// TIA Portal project "XSFW_TIA32701_A8" (V15.1)

(* hardware
DEVICE "S7-1200 station_1"  S7-1200 Station
   slot 0: "Rack_0"  S7-1200 Rack  Rack  V1.0
   slot 1: "PLC_1"  CPU 1212C DC/DC/DC  6ES7 212-1AE40-0XB0  V4.2
   slot 2: "DI 16/DQ 16x24VDC_1"  6ES7 223-1BL32-0XB0  V2.0
DEVICE "HMI_1"  KTP700 Basic PN
   slot 0: "HMI_1"  KTP700 Basic PN  6AV2 123-2GB03-0AX0  15.0.0.0
   slot 1: "HMI_RT_1"  KTP700 Basic PN  6AV2 123-2GB03-0AX0  15.0.0.0
   slot 5: "HMI_1.IE_CP_1"  PROFINET Interface  15.0.0.0
      slot 1: "Interfaz PROFINET_1"  PROFINET Interface
         slot 1: "Port_1"  Port
*)

// ===== PLC "PLC_1"  CPU 1212C DC/DC/DC =====

VAR_GLOBAL   // PLC tag table "Tabla de variables estándar"
   "Tag_2" AT %M101.0 : Bool;
   "Clock_Byte" AT %MB0 : Byte;
   "Clock_10Hz" AT %M0.0 : Bool;
   "Clock_5Hz" AT %M0.1 : Bool;
   "Clock_2.5Hz" AT %M0.2 : Bool;
   "Clock_2Hz" AT %M0.3 : Bool;
   "Clock_1.25Hz" AT %M0.4 : Bool;
   "Clock_1Hz" AT %M0.5 : Bool;
   "Clock_0.625Hz" AT %M0.6 : Bool;
   "Clock_0.5Hz" AT %M0.7 : Bool;
   "System_Byte" AT %MB1 : Byte;
   "FirstScan" AT %M1.0 : Bool;
   "DiagStatusUpdate" AT %M1.1 : Bool;
   "AlwaysTRUE" AT %M1.2 : Bool;
   "AlwaysFALSE" AT %M1.3 : Bool;
   "Alarma Activa" AT %M10.0 : Bool;   // Alarma Activa
   "Circuito_Seguridad" AT %M10.1 : Bool;   // circuito de seguridad
   "Tag_1" AT %M10.2 : Bool;
   "Marcha_Linea" AT %M127.4 : Bool;
   "Siempre 0" AT %M128.0 : Bool;
   "siempre 1" AT %M128.1 : Bool;
   "E0.0_FILT1segTensMand" AT %M128.2 : Bool;   // Filtracion de Tension de mando
   "clk_100ms" AT %M128.4 : Bool;
   "clk_1s" AT %M128.5 : Bool;   // clok de 1seg
   "clk_200ms" AT %M128.6 : Bool;   // clok 200ms
   "clk_350ms" AT %M128.7 : Bool;
   "Falla_rol_entra" AT %M129.1 : Bool;
   "clk_2s" AT %M129.6 : Bool;   // clok de 2seg
   "Tag_23" AT %M129.7 : Bool;
   "FALTA CONFIRMACION DE GUARDAM_rol_ent" AT %M160.1 : Bool;
   "Saturacion excesiva" AT %M160.5 : Bool;
   "Ord_Marc_Ord_Ent" AT %M160.7 : Bool;
   "En_ciclo" AT %M161.0 : Bool;   // En Ciclo
   "flipflop act/des FC6.7" AT %M161.1 : Bool;
   "Bajar_topeSolT" AT %M161.2 : Bool;   // bajar tope solapa trasero filtado TON
   "Ord_Disp_Cola" AT %M161.3 : Bool;
   "Sns_satur_ton" AT %M161.4 : Bool;   // Sensor de saturacion filtrado TON
   "E1.7_filtr_verificar" AT %M161.5 : Bool;   // E1.7 filtrado TON
   "Tag_3" AT %M300.0 : Bool;
   "Tag_4" AT %M200.0 : Bool;
   "Aux_Solapa_Abierta" AT %M2.4 : Bool;
END_VAR

VAR_GLOBAL   // PLC tag table "Entradas"
   "iTension_Mando" AT %E0.0 : Bool;   // Tension de mando
   "iParad_Emerg" AT %E0.1 : Bool;   // Pulsador parada de emergecia
   "iGmt_cin_later" AT %E0.3 : Bool;   // Guardamotor cintas laterales
   "iGmt_rolos_Ent" AT %E0.4 : Bool;   // Guardamotor rolos de entrada
   "iPls_Marcha" AT %E0.5 : Bool;   // pulsador de marcha
   "iPls_Parada" AT %E0.6 : Bool;   // pulsador de parada
   "iSel_Transf_Embalaje" AT %E0.7 : Bool;   // Selectora transferencia embalaje
   "iSel_Cola_Calien" AT %E1.0 : Bool;   // Selectora cola caliente
   "iSns_2Cin" AT %E1.1 : Bool;   // Sensor 2 cinta
   "iSns_3Cin" AT %E1.2 : Bool;   // Sensor 3 cinta
   "iSns_4Cin" AT %E1.3 : Bool;   // Sensor 4 cinta
   "iSns_5Cin" AT %E1.4 : Bool;   // Sensor 5 cinta
   "iSns_1Cin" AT %E1.5 : Bool;   // Sensor 1 cinta
   "iSns_Satur" AT %E1.6 : Bool;   // Sensor de saturacion
   "RELEVAR_SIEMP_LLEGA_1" AT %E1.7 : Bool;   // REVISAR siempre llega 1 Acum transp siguiente
   "iSns_Puerta_1" AT %E2.0 : Bool;   // Puerta 1
   "iSns_Puerta_2" AT %E2.1 : Bool;   // Puerta 2
   "iSns_Puerta_3" AT %E2.2 : Bool;   // Puerta 3
   "iSns_Puerta_4" AT %E2.3 : Bool;   // Puerta 4
   "iSns_Solapa_Abierta" AT %E2.4 : Bool;   // SOLAPA TRASERA ABIERTA
   "iReserva RESET I0.2" AT %I0.2 : Bool;   // Pulsador RESET
   "iReserva I2.5" AT %I2.5 : Bool;
   "iReserva I2.6" AT %I2.6 : Bool;
   "iReserva I2.7" AT %I2.7 : Bool;
END_VAR

VAR_GLOBAL   // PLC tag table "Salidas"
   "oCtc_Cin_Later" AT %A0.0 : Bool;   // Cintas Laterales
   "oCtc_Rod_Ent" AT %A0.1 : Bool;   // Rodillos de entrada
   "oCtc_Encolador" AT %A0.2 : Bool;   // Alim. encolador
   "oCil_Tope_solapa_Subir" AT %A0.3 : Bool;   // Levantar tope solapa
   "oDisp_Cola" AT %A0.4 : Bool;   // Bajar tope solapa trasera
   "oLmp_Falla" AT %A0.5 : Bool;   // Falla presente
   "oLmp__Marcha" AT %A1.0 : Bool;   // Testigo de marcha
   "oHab_Seguridades" AT %A1.1 : Bool;   // Habilita seguridades
   "oReserva A1.2" AT %Q1.2 : Bool;
   "oReserva A1.3" AT %Q1.3 : Bool;
   "oReserva A1.4" AT %Q1.4 : Bool;
   "oReserva A1.5" AT %Q1.5 : Bool;
   "oReserva A1.6" AT %Q1.6 : Bool;
   "oReserva A1.7" AT %Q1.7 : Bool;
   "oReserva A2.0" AT %Q2.0 : Bool;
   "oReserva A2.1" AT %Q2.1 : Bool;
   "oReserva A2.2" AT %Q2.2 : Bool;
   "oReserva A2.3" AT %Q2.3 : Bool;
   "oReserva A2.4" AT %Q2.4 : Bool;
   "oReserva A2.5" AT %Q2.5 : Bool;
   "oReserva A2.6" AT %Q2.6 : Bool;
   "oReserva A2.7" AT %Q2.7 : Bool;
END_VAR

DATA_BLOCK "DB1"   // DB1
{ S7_Optimized_Access := 'FALSE' }
VERSION : 0.0
   VAR
      D_0 : Word := WORD#16#4442;
      D_1 : Word := WORD#16#3120;
      D_2 : Word := WORD#16#4F42;
      D_3 : Word := WORD#16#413A;
      D_4 : Word := WORD#16#2041;
      D_5 : Word := WORD#16#4920;
      D_6 : Word := WORD#16#3020;
      D_7 : Word := WORD#16#3B20;
      D_8 : Word := WORD#16#4F42;
      D_9 : Word := WORD#16#493A;
      D_10 : Word := WORD#16#2020;
      D_11 : Word := WORD#16#2020;
      D_12 : Word := WORD#16#2020;
      D_13 : Word := WORD#16#203B;
      D_14 : Word := WORD#16#204F;
      D_15 : Word := WORD#16#4243;
      D_16 : Word := WORD#16#3A20;
      D_17 : Word := WORD#16#4341;
      D_18 : Word := WORD#16#5020;
      D_19 : Word := WORD#16#4E20;
      D_20 : Word := WORD#16#2020;
      D_21 : Word := WORD#16#2020;
      D_22 : Word := WORD#16#4342;
      D_23 : Word := WORD#16#5020;
      D_24 : Word := WORD#16#4E20;
      D_25 : Word := WORD#16#2020;
      D_26 : Word := WORD#16#2020;
      D_27 : Word := WORD#16#203B;
      D_28 : Word := WORD#16#2353;
      D_29 : Word := WORD#16#4C31;
      D_30 : Word := WORD#16#3A20;
      D_31 : Word := WORD#16#534C;
      D_32 : Word := WORD#16#4E20;
      D_33 : Word := WORD#16#3120;
      D_34 : Word := WORD#16#2053;
      D_35 : Word := WORD#16#4620;
      D_36 : Word := WORD#16#4442;
      D_37 : Word := WORD#16#3220;
      D_38 : Word := WORD#16#2044;
      D_39 : Word := WORD#16#5730;
      D_40 : Word := WORD#16#2020;
      D_41 : Word := WORD#16#2045;
      D_42 : Word := WORD#16#4620;
      D_43 : Word := WORD#16#4442;
      D_44 : Word := WORD#16#3320;
      D_45 : Word := WORD#16#2044;
      D_46 : Word := WORD#16#5730;
      D_47 : Word := WORD#16#2020;
      D_48 : Word := WORD#16#2020;
      D_49 : Word := WORD#16#4B42;
      D_50 : Word := WORD#16#4520;
      D_51 : Word := WORD#16#4D42;
      D_52 : Word := WORD#16#3130;
      D_53 : Word := WORD#16#3020;
      D_54 : Word := WORD#16#2020;
      D_55 : Word := WORD#16#2020;
      D_56 : Word := WORD#16#204B;
      D_57 : Word := WORD#16#4253;
      D_58 : Word := WORD#16#204D;
      D_59 : Word := WORD#16#4231;
      D_60 : Word := WORD#16#3031;
      D_61 : Word := WORD#16#2020;
      D_62 : Word := WORD#16#2020;
      D_63 : Word := WORD#16#2020;
      D_64 : Word := WORD#16#5047;
      D_65 : Word := WORD#16#4E20;
      D_66 : Word := WORD#16#3120;
      D_67 : Word := WORD#16#203B;
      D_68 : Word := WORD#16#2320;
      D_69 : Word := WORD#16#5344;
      D_70 : Word := WORD#16#503A;
      D_71 : Word := WORD#16#204E;
      D_72 : Word := WORD#16#5420;
      D_73 : Word := WORD#16#3132;
      D_74 : Word := WORD#16#3820;
      D_75 : Word := WORD#16#5042;
      D_76 : Word := WORD#16#5553;
      D_77 : Word := WORD#16#204E;
      D_78 : Word := WORD#16#203B;
      D_79 : Word := WORD#16#2054;
      D_80 : Word := WORD#16#4642;
      D_81 : Word := WORD#16#3A20;
      D_82 : Word := WORD#16#4F42;
      D_83 : Word := WORD#16#3133;
      D_84 : Word := WORD#16#2031;
      D_85 : Word := WORD#16#3030;
      D_86 : Word := WORD#16#2020;
      D_87 : Word := WORD#16#2020;
      D_88 : Word := WORD#16#3B20;
      D_89 : Word := WORD#16#2343;
      D_90 : Word := WORD#16#4C50;
      D_91 : Word := WORD#16#3A20;
      D_92 : Word := WORD#16#5354;
      D_93 : Word := WORD#16#5720;
      D_94 : Word := WORD#16#4D57;
      D_95 : Word := WORD#16#3130;
      D_96 : Word := WORD#16#3220;
      D_97 : Word := WORD#16#2020;
      D_98 : Word := WORD#16#2020;
      D_99 : Word := WORD#16#2020;
      D_100 : Word := WORD#16#2043;
      D_101 : Word := WORD#16#4C4B;
      D_102 : Word := WORD#16#2044;
      D_103 : Word := WORD#16#4235;
      D_104 : Word := WORD#16#2020;
      D_105 : Word := WORD#16#4457;
      D_106 : Word := WORD#16#3020;
      D_107 : Word := WORD#16#2020;
      D_108 : Word := WORD#16#2020;
      D_109 : Word := WORD#16#5345;
      D_110 : Word := WORD#16#5420;
      D_111 : Word := WORD#16#3320;
      D_112 : Word := WORD#16#2030;
      D_113 : Word := WORD#16#312E;
      D_114 : Word := WORD#16#3130;
      D_115 : Word := WORD#16#2E39;
      D_116 : Word := WORD#16#3120;
      D_117 : Word := WORD#16#3132;
      D_118 : Word := WORD#16#3A30;
      D_119 : Word := WORD#16#303A;
      D_120 : Word := WORD#16#3030;
      D_121 : Word := WORD#16#2020;
      D_122 : Word := WORD#16#2020;
      D_123 : Word := WORD#16#4F48;
      D_124 : Word := WORD#16#5320;
      D_125 : Word := WORD#16#3030;
      D_126 : Word := WORD#16#3030;
      D_127 : Word := WORD#16#3030;
      D_128 : Word := WORD#16#3A30;
      D_129 : Word := WORD#16#303A;
      D_130 : Word := WORD#16#3030;
      D_131 : Word := WORD#16#2020;
      D_132 : Word := WORD#16#2020;
      D_133 : Word := WORD#16#5449;
      D_134 : Word := WORD#16#5320;
      D_135 : Word := WORD#16#3320;
      D_136 : Word := WORD#16#3031;
      D_137 : Word := WORD#16#2E31;
      D_138 : Word := WORD#16#302E;
      D_139 : Word := WORD#16#2031;
      D_140 : Word := WORD#16#323A;
      D_141 : Word := WORD#16#3030;
      D_142 : Word := WORD#16#3A30;
      D_143 : Word := WORD#16#3020;
      D_144 : Word := WORD#16#2020;
      D_145 : Word := WORD#16#2053;
      D_146 : Word := WORD#16#5450;
      D_147 : Word := WORD#16#2059;
      D_148 : Word := WORD#16#2053;
      D_149 : Word := WORD#16#4156;
      D_150 : Word := WORD#16#2059;
      D_151 : Word := WORD#16#2020;
      D_152 : Word := WORD#16#4346;
      D_153 : Word := WORD#16#2030;
      D_154 : Word := WORD#16#3020;
      D_155 : Word := WORD#16#2020;
      D_156 : Word := WORD#16#203B;
      D_157 : Word := WORD#16#2023;
      D_158 : Word := WORD#16#454E;
      D_159 : Word := WORD#16#4420;
   END_VAR
BEGIN
END_DATA_BLOCK

DATA_BLOCK "Comandos"   // DB2
{ S7_Optimized_Access := 'TRUE' }
VERSION : 0.1
   VAR
      marcha_panel : Bool;
      parada_panel : Bool;
   END_VAR
BEGIN
END_DATA_BLOCK

DATA_BLOCK "HMI"   // DB3
{ S7_Optimized_Access := 'TRUE' }
VERSION : 0.1
   VAR RETAIN
      Tiem_Satur : Time := T#3s;
      Tiem_cicloCola : Time := T#800ms;
      Tiem_DisparoCola : Time := T#400ms;
   END_VAR
   VAR
      WAlarmas_1 : Word;
      RESET : Bool;
      Cartel_Pausa_Solapa : Bool;
      Cartel_Pausa_Saturación : Bool;
   END_VAR
   VAR RETAIN
      PAUSA_RODILLO_ENTRADA : Time := T#400ms;
   END_VAR
BEGIN
END_DATA_BLOCK

DATA_BLOCK "Temporizadores"   // DB11
{ S7_Optimized_Access := 'TRUE' }
VERSION : 0.1
   VAR RETAIN
      T1 : IEC_TIMER;
      T2 : IEC_TIMER;
      T3 : IEC_TIMER;
      T4 : IEC_TIMER;
      T5 : IEC_TIMER;
      T6 : IEC_TIMER;
      T7 : IEC_TIMER;
      T8 : IEC_TIMER;
      T9 : IEC_TIMER;
      T10 : IEC_TIMER;
      T11 : IEC_TIMER;
      T12 : IEC_TIMER;
      T13 : IEC_TIMER;
      T14 : IEC_TIMER;
      T15 : IEC_TIMER;
      T16 : IEC_TIMER;
      T17 : IEC_TIMER;
      T18 : IEC_TIMER;
      T19 : IEC_TIMER;
      T20 : IEC_TIMER;
      T21 : IEC_TIMER;
      T22 : IEC_TIMER;
      T23 : IEC_TIMER;
      T24 : IEC_TIMER;
      T25 : IEC_TIMER;
      T26 : IEC_TIMER;
      T27 : IEC_TIMER;
      T28 : IEC_TIMER;
      T29 : IEC_TIMER;
      T30 : IEC_TIMER;
      T31 : IEC_TIMER;
      T32 : IEC_TIMER;
      Tiempo1 : Time := T#2s;
      Tiempo2 : Time;
      Tiempo3 : Time;
      Tiempo4 : Time;
      Tiempo5 : Time;
      Tiempo6 : Time;
      Tiempo7 : Time;
      Tiempo8 : Time;
      Tiempo9 : Time;
      Tiempo10 : Time;
      Tiempo11 : Time;
      Tiempo12 : Time;
      Tiempo13 : Time;
      Tiempo14 : Time;
      Tiempo15 : Time;
      Tiempo16 : Time;
      Tiempo17 : Time;
      Tiempo18 : Time;
      Tiempo19 : Time;
      Tiempo20 : Time;
      Tiempo21 : Time;
      Tiempo22 : Time;
      Tiempo23 : Time;
      Tiempo24 : Time;
      Tiempo25 : Time;
      Tiempo26 : Time;
      Tiempo27 : Time;
      Tiempo28 : Time;
      Tiempo29 : Time;
      Tiempo30 : Time;
      Tiempo31 : Time;
      Tiempo32 : Time;
   END_VAR
BEGIN
END_DATA_BLOCK

// folder: System blocks/Program resources

DATA_BLOCK "Filtr1s"   // DB4
{ S7_Optimized_Access := 'TRUE' }
AUTHOR : Simatic
FAMILY : IEC
NAME : IEC_TMR
VERSION : 1.0
// stored: InstanceOfName IEC_TIMER
"IEC_TIMER"
BEGIN
END_DATA_BLOCK

DATA_BLOCK "IEC_Timer_0_DB"   // DB5
{ S7_Optimized_Access := 'TRUE' }
AUTHOR : Simatic
FAMILY : IEC
NAME : IEC_TMR
VERSION : 1.0
// stored: InstanceOfName IEC_TIMER
"IEC_TIMER"
BEGIN
END_DATA_BLOCK

DATA_BLOCK "ta_11"   // DB7
{ S7_Optimized_Access := 'TRUE' }
AUTHOR : Simatic
FAMILY : IEC
NAME : IEC_TMR
VERSION : 1.0
// stored: InstanceOfName IEC_TIMER
"IEC_TIMER"
BEGIN
END_DATA_BLOCK

DATA_BLOCK "ta_13"   // DB8
{ S7_Optimized_Access := 'TRUE' }
AUTHOR : Simatic
FAMILY : IEC
NAME : IEC_TMR
VERSION : 1.0
// stored: InstanceOfName IEC_TIMER
"IEC_TIMER"
BEGIN
END_DATA_BLOCK

DATA_BLOCK "ton sensor saturacion"   // DB9
{ S7_Optimized_Access := 'TRUE' }
AUTHOR : Simatic
FAMILY : IEC
NAME : IEC_TMR
VERSION : 1.0
// stored: InstanceOfName IEC_TIMER
"IEC_TIMER"
BEGIN
END_DATA_BLOCK

DATA_BLOCK "ta_51"   // DB10
{ S7_Optimized_Access := 'TRUE' }
AUTHOR : Simatic
FAMILY : IEC
NAME : IEC_TMR
VERSION : 1.0
// stored: InstanceOfName IEC_TIMER
"IEC_TIMER"
BEGIN
END_DATA_BLOCK

DATA_BLOCK "TON DE 1s - E1.5 Sns_1Cin"   // DB12
{ S7_Optimized_Access := 'TRUE' }
AUTHOR : Simatic
FAMILY : IEC
NAME : IEC_TMR
VERSION : 1.0
// stored: InstanceOfName IEC_TIMER
"IEC_TIMER"
BEGIN
END_DATA_BLOCK

DATA_BLOCK "IEC_Timer_0_DB_1"   // DB13
{ S7_Optimized_Access := 'TRUE' }
AUTHOR : Simatic
FAMILY : IEC
NAME : IEC_TMR
VERSION : 1.0
// stored: InstanceOfName IEC_TIMER
"IEC_TIMER"
BEGIN
END_DATA_BLOCK

DATA_BLOCK "TON 5s rolos_entra_ funcionamiento"   // DB14
{ S7_Optimized_Access := 'TRUE' }
AUTHOR : Simatic
FAMILY : IEC
NAME : IEC_TMR
VERSION : 1.0
// stored: InstanceOfName IEC_TIMER
"IEC_TIMER"
BEGIN
END_DATA_BLOCK

DATA_BLOCK "ta_71"   // DB15
{ S7_Optimized_Access := 'TRUE' }
AUTHOR : Simatic
FAMILY : IEC
NAME : IEC_TMR
VERSION : 1.0
// stored: InstanceOfName IEC_TIMER
"IEC_TIMER"
BEGIN
END_DATA_BLOCK

DATA_BLOCK "PAUSA_SATUR"   // DB18
{ S7_Optimized_Access := 'TRUE' }
AUTHOR : Simatic
FAMILY : IEC
NAME : IEC_TMR
VERSION : 1.0
// stored: InstanceOfName IEC_TIMER
"IEC_TIMER"
BEGIN
END_DATA_BLOCK

DATA_BLOCK "ta_15"   // DB19
{ S7_Optimized_Access := 'TRUE' }
AUTHOR : Simatic
FAMILY : IEC
NAME : IEC_TMR
VERSION : 1.0
// stored: InstanceOfName IEC_TIMER
"IEC_TIMER"
BEGIN
END_DATA_BLOCK

DATA_BLOCK "ta_16"   // DB20
{ S7_Optimized_Access := 'TRUE' }
AUTHOR : Simatic
FAMILY : IEC
NAME : IEC_TMR
VERSION : 1.0
// stored: InstanceOfName IEC_TIMER
"IEC_TIMER"
BEGIN
END_DATA_BLOCK

DATA_BLOCK "ta_18"   // DB21
{ S7_Optimized_Access := 'TRUE' }
AUTHOR : Simatic
FAMILY : IEC
NAME : IEC_TMR
VERSION : 1.0
// stored: InstanceOfName IEC_TIMER
"IEC_TIMER"
BEGIN
END_DATA_BLOCK

DATA_BLOCK "ta_19"   // DB22
{ S7_Optimized_Access := 'TRUE' }
AUTHOR : Simatic
FAMILY : IEC
NAME : IEC_TMR
VERSION : 1.0
// stored: InstanceOfName IEC_TIMER
"IEC_TIMER"
BEGIN
END_DATA_BLOCK

DATA_BLOCK "ta_21"   // DB23
{ S7_Optimized_Access := 'TRUE' }
AUTHOR : Simatic
FAMILY : IEC
NAME : IEC_TMR
VERSION : 1.0
// stored: InstanceOfName IEC_TIMER
"IEC_TIMER"
BEGIN
END_DATA_BLOCK

DATA_BLOCK "ta_22"   // DB24
{ S7_Optimized_Access := 'TRUE' }
AUTHOR : Simatic
FAMILY : IEC
NAME : IEC_TMR
VERSION : 1.0
// stored: InstanceOfName IEC_TIMER
"IEC_TIMER"
BEGIN
END_DATA_BLOCK

// folder: (top level)

FUNCTION "Alarmas" : Void   // FC1, LAD
{ S7_Optimized_Access := 'TRUE' }
VERSION : 0.1
BEGIN

REGION Network 1: FALLA ACTIVA EN CIRCUITO DE SEGURIDAD
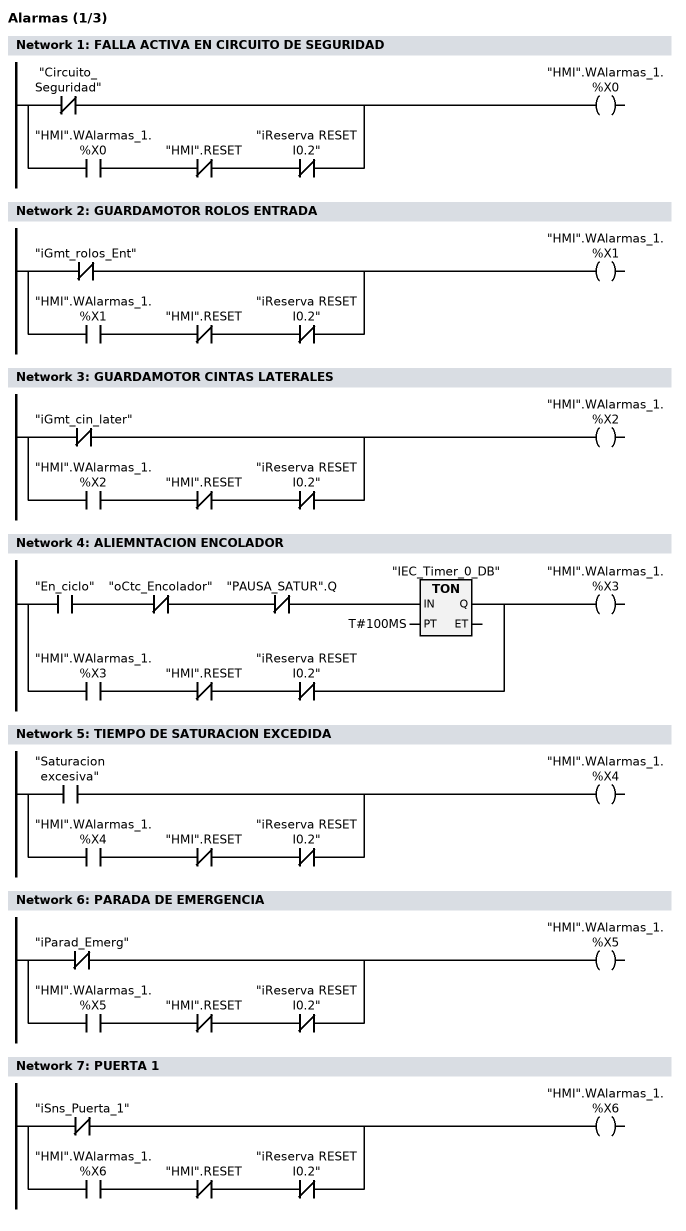
   RUNG wire#powerrail
      I_Contact( "Circuito_Seguridad" )
      wire#w1
      Coil( "HMI".WAlarmas_1.%X0 )
   END_RUNG
   RUNG wire#powerrail
      Contact( "HMI".WAlarmas_1.%X0 )
      I_Contact( "HMI".RESET )
      I_Contact( "iReserva RESET I0.2" )
   END_RUNG wire#w1
   // the same network as SCL:
   "HMI".WAlarmas_1.%X0 := NOT "Circuito_Seguridad" OR ("HMI".WAlarmas_1.%X0 AND NOT "HMI".RESET AND NOT "iReserva RESET I0.2");
END_REGION

REGION Network 2: GUARDAMOTOR ROLOS ENTRADA
   RUNG wire#powerrail
      I_Contact( "iGmt_rolos_Ent" )
      wire#w1
      Coil( "HMI".WAlarmas_1.%X1 )
   END_RUNG
   RUNG wire#powerrail
      Contact( "HMI".WAlarmas_1.%X1 )
      I_Contact( "HMI".RESET )
      I_Contact( "iReserva RESET I0.2" )
   END_RUNG wire#w1
   // the same network as SCL:
   "HMI".WAlarmas_1.%X1 := NOT "iGmt_rolos_Ent" OR ("HMI".WAlarmas_1.%X1 AND NOT "HMI".RESET AND NOT "iReserva RESET I0.2");
END_REGION

REGION Network 3: GUARDAMOTOR CINTAS LATERALES
   RUNG wire#powerrail
      I_Contact( "iGmt_cin_later" )
      wire#w1
      Coil( "HMI".WAlarmas_1.%X2 )
   END_RUNG
   RUNG wire#powerrail
      Contact( "HMI".WAlarmas_1.%X2 )
      I_Contact( "HMI".RESET )
      I_Contact( "iReserva RESET I0.2" )
   END_RUNG wire#w1
   // the same network as SCL:
   "HMI".WAlarmas_1.%X2 := NOT "iGmt_cin_later" OR ("HMI".WAlarmas_1.%X2 AND NOT "HMI".RESET AND NOT "iReserva RESET I0.2");
END_REGION

REGION Network 4: ALIEMNTACION ENCOLADOR
   "IEC_Timer_0_DB".TON(IN := "En_ciclo" AND NOT "oCtc_Encolador" AND NOT "PAUSA_SATUR".Q, PT := T#100MS);
   "HMI".WAlarmas_1.%X3 := "IEC_Timer_0_DB".Q OR ("HMI".WAlarmas_1.%X3 AND NOT "HMI".RESET AND NOT "iReserva RESET I0.2");
END_REGION

REGION Network 5: TIEMPO DE SATURACION EXCEDIDA
   RUNG wire#powerrail
      Contact( "Saturacion excesiva" )
      wire#w1
      Coil( "HMI".WAlarmas_1.%X4 )
   END_RUNG
   RUNG wire#powerrail
      Contact( "HMI".WAlarmas_1.%X4 )
      I_Contact( "HMI".RESET )
      I_Contact( "iReserva RESET I0.2" )
   END_RUNG wire#w1
   // the same network as SCL:
   "HMI".WAlarmas_1.%X4 := "Saturacion excesiva" OR ("HMI".WAlarmas_1.%X4 AND NOT "HMI".RESET AND NOT "iReserva RESET I0.2");
END_REGION

REGION Network 6: PARADA DE EMERGENCIA
   RUNG wire#powerrail
      I_Contact( "iParad_Emerg" )
      wire#w1
      Coil( "HMI".WAlarmas_1.%X5 )
   END_RUNG
   RUNG wire#powerrail
      Contact( "HMI".WAlarmas_1.%X5 )
      I_Contact( "HMI".RESET )
      I_Contact( "iReserva RESET I0.2" )
   END_RUNG wire#w1
   // the same network as SCL:
   "HMI".WAlarmas_1.%X5 := NOT "iParad_Emerg" OR ("HMI".WAlarmas_1.%X5 AND NOT "HMI".RESET AND NOT "iReserva RESET I0.2");
END_REGION

REGION Network 7: PUERTA 1
   RUNG wire#powerrail
      I_Contact( "iSns_Puerta_1" )
      wire#w1
      Coil( "HMI".WAlarmas_1.%X6 )
   END_RUNG
   RUNG wire#powerrail
      Contact( "HMI".WAlarmas_1.%X6 )
      I_Contact( "HMI".RESET )
      I_Contact( "iReserva RESET I0.2" )
   END_RUNG wire#w1
   // the same network as SCL:
   "HMI".WAlarmas_1.%X6 := NOT "iSns_Puerta_1" OR ("HMI".WAlarmas_1.%X6 AND NOT "HMI".RESET AND NOT "iReserva RESET I0.2");
END_REGION

REGION Network 8: PUERTA 2
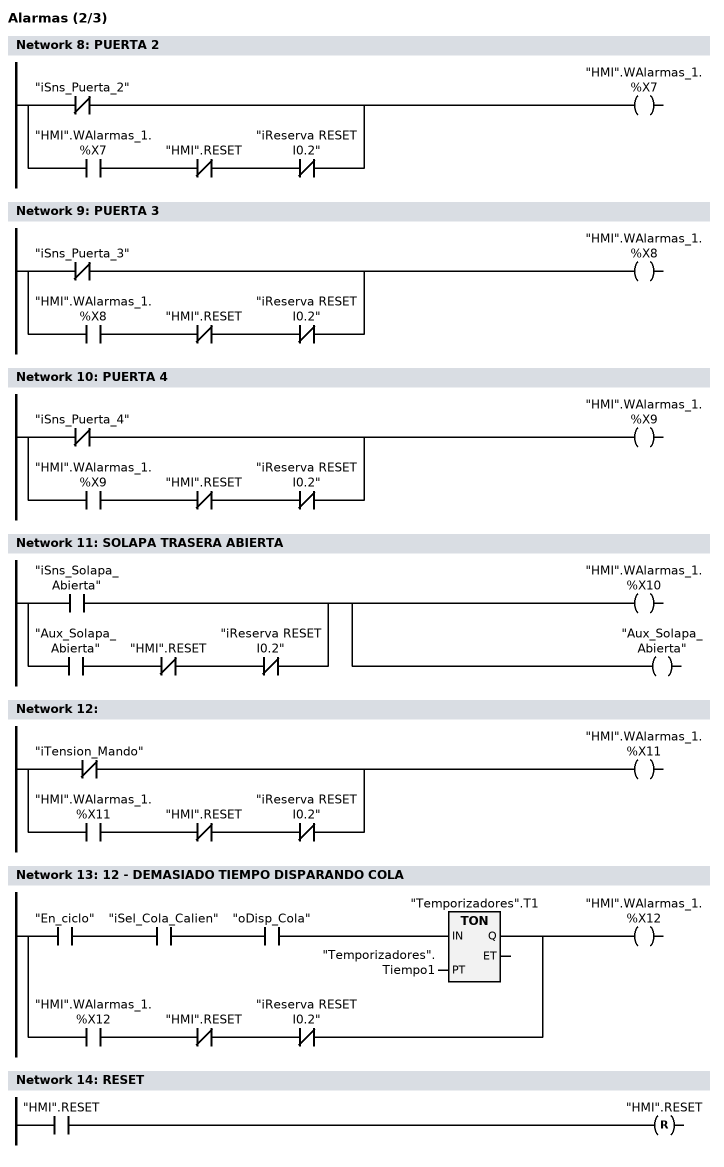
   RUNG wire#powerrail
      I_Contact( "iSns_Puerta_2" )
      wire#w1
      Coil( "HMI".WAlarmas_1.%X7 )
   END_RUNG
   RUNG wire#powerrail
      Contact( "HMI".WAlarmas_1.%X7 )
      I_Contact( "HMI".RESET )
      I_Contact( "iReserva RESET I0.2" )
   END_RUNG wire#w1
   // the same network as SCL:
   "HMI".WAlarmas_1.%X7 := NOT "iSns_Puerta_2" OR ("HMI".WAlarmas_1.%X7 AND NOT "HMI".RESET AND NOT "iReserva RESET I0.2");
END_REGION

REGION Network 9: PUERTA 3
   RUNG wire#powerrail
      I_Contact( "iSns_Puerta_3" )
      wire#w1
      Coil( "HMI".WAlarmas_1.%X8 )
   END_RUNG
   RUNG wire#powerrail
      Contact( "HMI".WAlarmas_1.%X8 )
      I_Contact( "HMI".RESET )
      I_Contact( "iReserva RESET I0.2" )
   END_RUNG wire#w1
   // the same network as SCL:
   "HMI".WAlarmas_1.%X8 := NOT "iSns_Puerta_3" OR ("HMI".WAlarmas_1.%X8 AND NOT "HMI".RESET AND NOT "iReserva RESET I0.2");
END_REGION

REGION Network 10: PUERTA 4
   RUNG wire#powerrail
      I_Contact( "iSns_Puerta_4" )
      wire#w1
      Coil( "HMI".WAlarmas_1.%X9 )
   END_RUNG
   RUNG wire#powerrail
      Contact( "HMI".WAlarmas_1.%X9 )
      I_Contact( "HMI".RESET )
      I_Contact( "iReserva RESET I0.2" )
   END_RUNG wire#w1
   // the same network as SCL:
   "HMI".WAlarmas_1.%X9 := NOT "iSns_Puerta_4" OR ("HMI".WAlarmas_1.%X9 AND NOT "HMI".RESET AND NOT "iReserva RESET I0.2");
END_REGION

REGION Network 11: SOLAPA TRASERA ABIERTA
   RUNG wire#powerrail
      Contact( "iSns_Solapa_Abierta" )
      wire#w1
      Coil( "HMI".WAlarmas_1.%X10 )
   END_RUNG
   RUNG wire#powerrail
      Contact( "Aux_Solapa_Abierta" )
      I_Contact( "HMI".RESET )
      I_Contact( "iReserva RESET I0.2" )
   END_RUNG wire#w1
   RUNG wire#w1
      Coil( "Aux_Solapa_Abierta" )
   END_RUNG
   // the same network as SCL:
   "HMI".WAlarmas_1.%X10 := "iSns_Solapa_Abierta" OR ("Aux_Solapa_Abierta" AND NOT "HMI".RESET AND NOT "iReserva RESET I0.2");
   "Aux_Solapa_Abierta" := "HMI".WAlarmas_1.%X10;
END_REGION

REGION Network 12
   RUNG wire#powerrail
      I_Contact( "iTension_Mando" )
      wire#w1
      Coil( "HMI".WAlarmas_1.%X11 )
   END_RUNG
   RUNG wire#powerrail
      Contact( "HMI".WAlarmas_1.%X11 )
      I_Contact( "HMI".RESET )
      I_Contact( "iReserva RESET I0.2" )
   END_RUNG wire#w1
   // the same network as SCL:
   "HMI".WAlarmas_1.%X11 := NOT "iTension_Mando" OR ("HMI".WAlarmas_1.%X11 AND NOT "HMI".RESET AND NOT "iReserva RESET I0.2");
END_REGION

REGION Network 13: 12 - DEMASIADO TIEMPO DISPARANDO COLA
   "Temporizadores".T1.TON(IN := "En_ciclo" AND "iSel_Cola_Calien" AND "oDisp_Cola",
                           PT := "Temporizadores".Tiempo1);
   "HMI".WAlarmas_1.%X12 := "Temporizadores".T1.Q OR ("HMI".WAlarmas_1.%X12 AND NOT "HMI".RESET AND NOT "iReserva RESET I0.2");
END_REGION

REGION Network 14: RESET
   RUNG wire#powerrail
      Contact( "HMI".RESET )
      R_Coil( "HMI".RESET )
   END_RUNG
   // the same network as SCL:
   IF "HMI".RESET THEN "HMI".RESET := FALSE; END_IF;
END_REGION

REGION Network 15: Alarma Activa
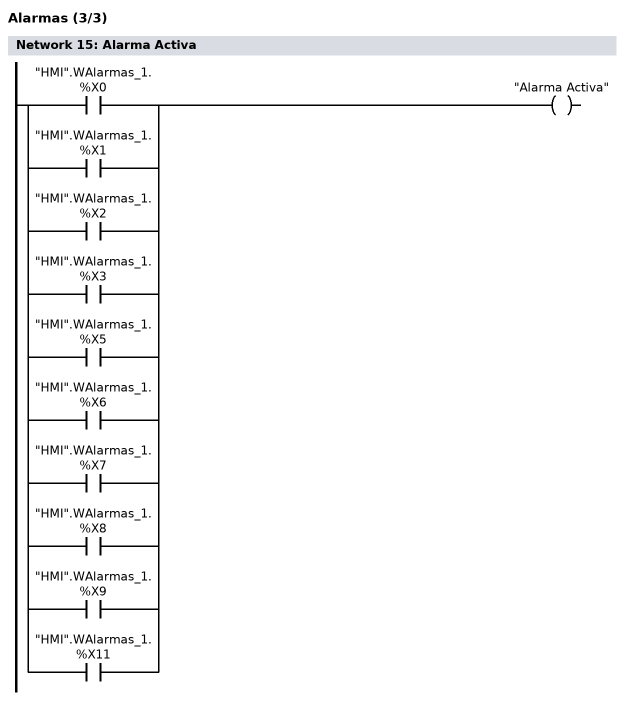
   RUNG wire#powerrail
      Contact( "HMI".WAlarmas_1.%X0 )
      wire#w1
      Coil( "Alarma Activa" )
   END_RUNG
   RUNG wire#powerrail
      Contact( "HMI".WAlarmas_1.%X1 )
   END_RUNG wire#w1
   RUNG wire#powerrail
      Contact( "HMI".WAlarmas_1.%X2 )
   END_RUNG wire#w1
   RUNG wire#powerrail
      Contact( "HMI".WAlarmas_1.%X3 )
   END_RUNG wire#w1
   RUNG wire#powerrail
      Contact( "HMI".WAlarmas_1.%X5 )
   END_RUNG wire#w1
   RUNG wire#powerrail
      Contact( "HMI".WAlarmas_1.%X6 )
   END_RUNG wire#w1
   RUNG wire#powerrail
      Contact( "HMI".WAlarmas_1.%X7 )
   END_RUNG wire#w1
   RUNG wire#powerrail
      Contact( "HMI".WAlarmas_1.%X8 )
   END_RUNG wire#w1
   RUNG wire#powerrail
      Contact( "HMI".WAlarmas_1.%X9 )
   END_RUNG wire#w1
   RUNG wire#powerrail
      Contact( "HMI".WAlarmas_1.%X11 )
   END_RUNG wire#w1
   // the same network as SCL:
   "Alarma Activa" := "HMI".WAlarmas_1.%X0 OR "HMI".WAlarmas_1.%X1 OR "HMI".WAlarmas_1.%X2 OR "HMI".WAlarmas_1.%X3 OR "HMI".WAlarmas_1.%X5 OR "HMI".WAlarmas_1.%X6 OR "HMI".WAlarmas_1.%X7 OR "HMI".WAlarmas_1.%X8 OR "HMI".WAlarmas_1.%X9 OR "HMI".WAlarmas_1.%X11;
END_REGION
END_FUNCTION

FUNCTION "Marcas de Sistema" : Void   // FC2, LAD
{ S7_Optimized_Access := 'TRUE' }
VERSION : 0.1
   VAR_TEMP   // added for the SCL form of the ladder/FBD networks
      _w1 : Bool;
   END_VAR
BEGIN

REGION Network 1: variable siempre 0 y 1
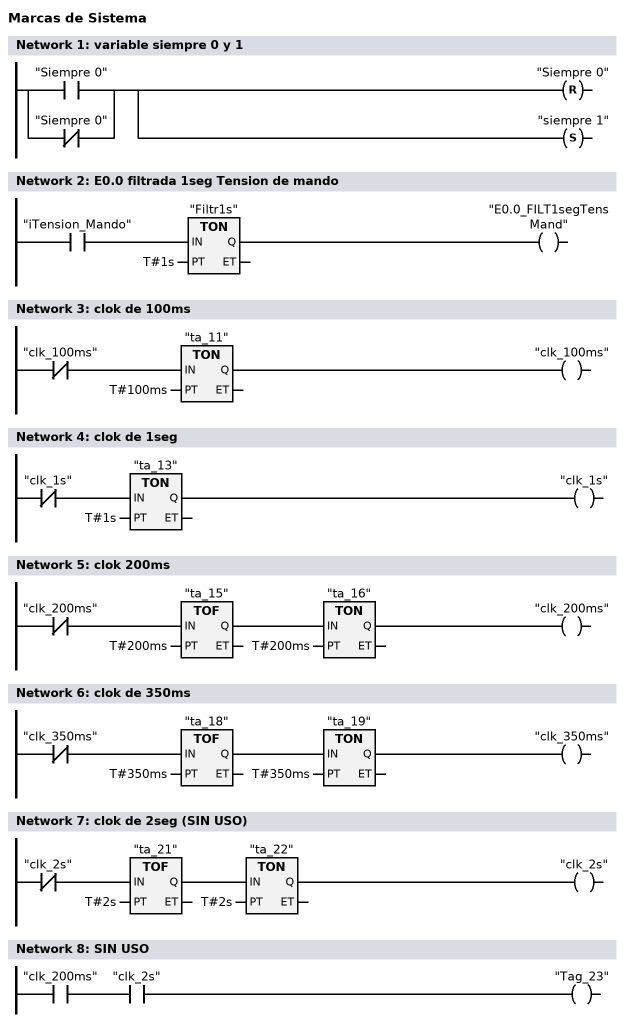
   RUNG wire#powerrail
      Contact( "Siempre 0" )
      wire#w1
      R_Coil( "Siempre 0" )
   END_RUNG
   RUNG wire#powerrail
      I_Contact( "Siempre 0" )
   END_RUNG wire#w1
   RUNG wire#w1
      S_Coil( "siempre 1" )
   END_RUNG
   // the same network as SCL:
   #_w1 := "Siempre 0" OR NOT "Siempre 0";
   IF #_w1 THEN
       "Siempre 0" := FALSE;
       "siempre 1" := TRUE;
   END_IF;
END_REGION

REGION Network 2: E0.0 filtrada 1seg Tension de mando
   "Filtr1s".TON(IN := "iTension_Mando", PT := T#1s);
   "E0.0_FILT1segTensMand" := "Filtr1s".Q;
END_REGION

REGION Network 3: clok de 100ms
   "ta_11".TON(IN := NOT "clk_100ms", PT := T#100ms);
   "clk_100ms" := "ta_11".Q;
END_REGION

REGION Network 4: clok de 1seg
   "ta_13".TON(IN := NOT "clk_1s", PT := T#1s);
   "clk_1s" := "ta_13".Q;
END_REGION

REGION Network 5: clok 200ms
   "ta_15".TOF(IN := NOT "clk_200ms", PT := T#200ms);
   "ta_16".TON(IN := "ta_15".Q, PT := T#200ms);
   "clk_200ms" := "ta_16".Q;
END_REGION

REGION Network 6: clok de 350ms
   "ta_18".TOF(IN := NOT "clk_350ms", PT := T#350ms);
   "ta_19".TON(IN := "ta_18".Q, PT := T#350ms);
   "clk_350ms" := "ta_19".Q;
END_REGION

REGION Network 7: clok de 2seg (SIN USO)
   "ta_21".TOF(IN := NOT "clk_2s", PT := T#2s);
   "ta_22".TON(IN := "ta_21".Q, PT := T#2s);
   "clk_2s" := "ta_22".Q;
END_REGION

REGION Network 8: SIN USO
   RUNG wire#powerrail
      Contact( "clk_200ms" )
      Contact( "clk_2s" )
      Coil( "Tag_23" )
   END_RUNG
   // the same network as SCL:
   "Tag_23" := "clk_200ms" AND "clk_2s";
END_REGION
END_FUNCTION

FUNCTION "FC6" : Void   // FC6, LAD
{ S7_Optimized_Access := 'TRUE' }
VERSION : 0.1
   VAR_TEMP
      Aux_TiempoDisp : Time;
   END_VAR
   VAR_TEMP   // added for the SCL form of the ladder/FBD networks
      _w1 : Bool;
   END_VAR
BEGIN

REGION Network 1: circuito de seguridad
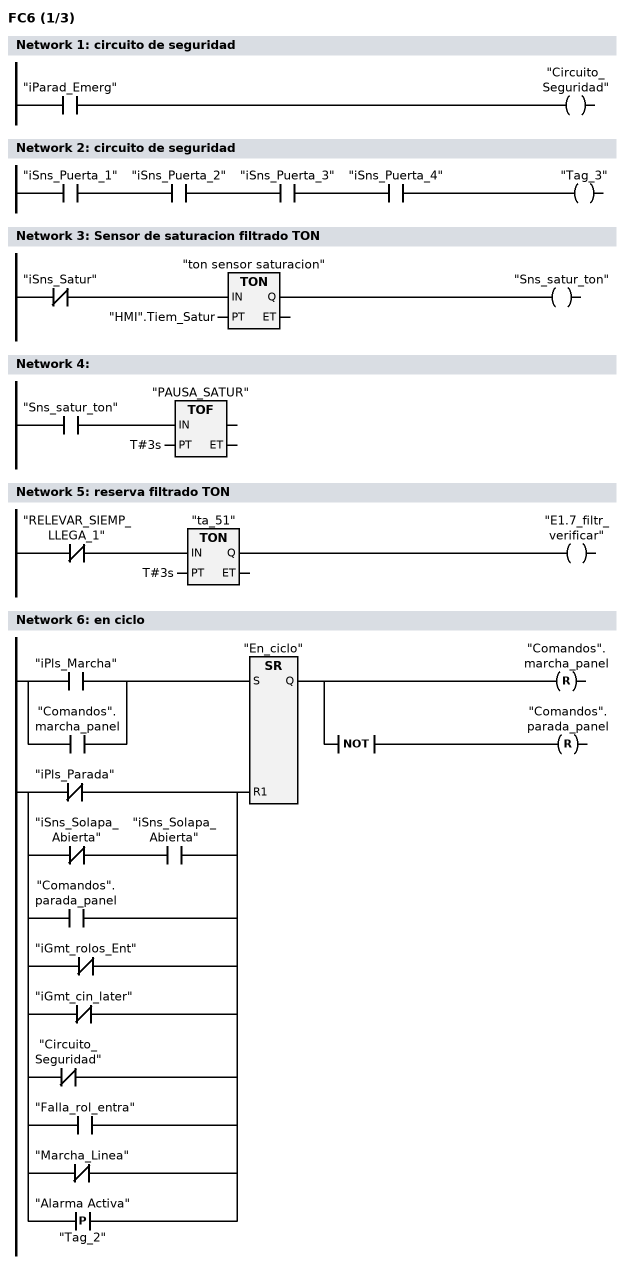
   RUNG wire#powerrail
      Contact( "iParad_Emerg" )
      Coil( "Circuito_Seguridad" )
   END_RUNG
   // the same network as SCL:
   "Circuito_Seguridad" := "iParad_Emerg";
END_REGION

REGION Network 2: circuito de seguridad
   RUNG wire#powerrail
      Contact( "iSns_Puerta_1" )
      Contact( "iSns_Puerta_2" )
      Contact( "iSns_Puerta_3" )
      Contact( "iSns_Puerta_4" )
      Coil( "Tag_3" )
   END_RUNG
   // the same network as SCL:
   "Tag_3" := "iSns_Puerta_1" AND "iSns_Puerta_2" AND "iSns_Puerta_3" AND "iSns_Puerta_4";
END_REGION

REGION Network 3: Sensor de saturacion filtrado TON
   "ton sensor saturacion".TON(IN := NOT "iSns_Satur", PT := "HMI".Tiem_Satur);
   "Sns_satur_ton" := "ton sensor saturacion".Q;
END_REGION

REGION Network 4
   "PAUSA_SATUR".TOF(IN := "Sns_satur_ton", PT := T#3s);
END_REGION

REGION Network 5: reserva filtrado TON
   "ta_51".TON(IN := NOT "RELEVAR_SIEMP_LLEGA_1", PT := T#3s);
   "E1.7_filtr_verificar" := "ta_51".Q;
END_REGION
